 '~Spare WB1[63].6'; 2023 '~Spare WB1[63].7'; 2024 '~Spare WB1[63].8'; 2025 '~Spare WB1[63].9'; 2026 '~Spare WB1[63].10'; 2027 '~Spare WB1[63].11'; 2028 '~Spare WB1[63].12'; 2029 '~Spare WB1[63].13'; 2030 '~Spare WB1[63].14'; 2031 '~Spare WB1[63].15'; 2032 '~Spare WB1[63].16'; 2033 '~Spare WB1[63].17'; 2034 '~Spare WB1[63].18'; 2035 '~Spare WB1[63].19'; 2036 '~Spare WB1[63].20'; 2037 '~Spare WB1[63].21'; 2038 '~Spare WB1[63].22'; 2039 '~Spare WB1[63].23'; 2040 '~Spare WB1[63].24'; 2041 '~Spare WB1[63].25'; 2042 '~Spare WB1[63].26'; 2043 '~Spare WB1[63].27'; 2044 '~Spare WB1[63].28'; 2045 '~Spare WB1[63].29'; 2046 '~Spare WB1[63].30'; 2047 '~Spare WB1[63].31'; 2048 '~Spare WB1[64].0'; 2049 '~Spare WB1[64].1'; 2050 '~Spare WB1[64].2'; 2051 '~Spare WB1[64].3'; 2052 '~Spare WB1[64].4'; 2053 '~Spare WB1[64].5'; 2054 '~Spare WB1[64].6'; 2055 '~Spare WB1[64].7'; 2056 '~Spare WB1[64].8'; 2057 '~Spare WB1[64].9'; 2058 '~Spare WB1[64].10'; 2059 '~Spare WB1[64].11'; 2060 '~Spare WB1[64].12'; 2061 '~Spare WB1[64].13'; 2062 '~Spare WB1[64].14'; 2063 '~Spare WB1[64].15'; 2064 '~Spare WB1[64].16'; 2065 '~Spare WB1[64].17'; 2066 '~Spare WB1[64].18'; 2067 '~Spare WB1[64].19'; 2068 '~Spare WB1[64].20'; 2069 '~Spare WB1[64].21'; 2070 '~Spare WB1[64].22'; 2071 '~Spare WB1[64].23'; 2072 '~Spare WB1[64].24'; 2073 '~Spare WB1[64].25'; 2074 '~Spare WB1[64].26'; 2075 '~Spare WB1[64].27'; 2076 '~Spare WB1[64].28'; 2077 '~Spare WB1[64].29'; 2078 '~Spare WB1[64].30'; 2079 '~Spare WB1[64].31'; 2080 '~Spare WB1[65].0'; 2081 '~Spare WB1[65].1'; 2082 '~Spare WB1[65].2'; 2083 '~Spare WB1[65].3'; 2084 '~Spare WB1[65].4'; 2085 '~Spare WB1[65].5'; 2086 '~Spare WB1[65].6'; 2087 '~Spare WB1[65].7'; 2088 '~Spare WB1[65].8'; 2089 '~Spare WB1[65].9'; 2090 '~Spare WB1[65].10'; 2091 '~Spare WB1[65].11'; 2092 '~Spare WB1[65].12'; 2093 '~Spare WB1[65].13'; 2094 '~Spare WB1[65].14'; 2095 '~Spare WB1[65].15'; 2096 '~Spare WB1[65].16'; 2097 '~Spare WB1[65].17'; 2098 '~Spare WB1[65].18'; 2099 '~Spare WB1[65].19'; 2100 '~Spare WB1[65].20'; 2101 '~Spare WB1[65].21'; 2102 '~Spare WB1[65].22'; 2103 '~Spare WB1[65].23'; 2104 '~Spare WB1[65].24'; 2105 '~Spare WB1[65].25'; 2106 '~Spare WB1[65].26'; 2107 '~Spare WB1[65].27'; 2108 '~Spare WB1[65].28'; 2109 '~Spare WB1[65].29'; 2110 '~Spare WB1[65].30'; 2111 '~Spare WB1[65].31'; 2112 '~S001R08 Waiting Zone #1 Not Clear WB1[66].0'; 2113 '~S001R08 Waiting Zone #2 Not Clear WB1[66].1'; 2114 '~S001R08 Waiting Zone #3 Not Clear WB1[66].2'; 2115 '~S001R08 Waiting Zone #4 Not Clear WB1[66].3'; 2116 '~S001R08 Waiting Zone #5 Not Clear WB1[66].4'; 2117 '~S001R08 Waiting Zone #6 Not Clear WB1[66].5'; 2118 '~S001R08 Waiting Zone #7 Not Clear WB1[66].6'; 2119 '~S001R08 Waiting Zone #8 Not Clear WB1[66].7'; 2120 '~S001R08 Waiting Zone #9 Not Clear WB1[66].8'; 2121 '~S001R08 Waiting Zone #10 Not Clear WB1[66].9'; 2122 '~S001R08 Waiting Zone #11 Not Clear WB1[66].10'; 2123 '~S001R08 Waiting Zone #12 Not Clear WB1[66].11'; 2124 '~S001R08 Waiting Zone #13 Not Clear WB1[66].12'; 2125 '~S001R08 Waiting Zone #14 Not Clear WB1[66].13'; 2126 '~S001R08 Waiting Tip Dress Zone #1 Not Clear WB1[66].14'; 2127 '~S001R08 Waiting Tip Dress Zone #2 Not Clear WB1[66].15'; 2128 '~S001R08 Adjacent Robot xx-xx In Teach WB1[66].16'; 2129 '~S001R08 Adjacent Robot xx-xx In Teach WB1[66].17'; 2130 '~S001R08 Adjacent Robot xx-xx In Teach WB1[66].18'; 2131 '~S001R08 Adjacent Robot xx-xx In Teach WB1[66].19'; 2132 '~S001R08 Adjacent Robot xx-xx In Teach WB1[66].20'; 2133 '~S001R08 Adjacent Robot xx-xx In Teach WB1[66].21'; 2134 '~S001R08 Adjacent Robot xx-xx In Teach WB1[66].22'; 2135 '~S001R08 Adjacent Robot xx-xx In Teach WB1[66].23'; 2136 '~S001R08 Adjacent Robot xx-xx In Teach WB1[66].24'; 2137 '~S001R08 Adjacent Robot xx-xx In Teach WB1[66].25'; 2138 '~Spare WB1[66].26'; 2139 '~Spare WB1[66].27'; 2140 '~Spare WB1[66].28'; 2141 '~S001R08 Robot Not Clear Of Fixture WB1[66].29'; 2142 '~Spare WB1[66].30'; 2143 '~Spare WB1[66].31'; 2144 '~Spare WB1[67].0'; 2145 '~Spare WB1[67].1'; 2146 '~Spare WB1[67].2'; 2147 '~Spare WB1[67].3'; 2148 '~Spare WB1[67].4'; 2149 '~Spare WB1[67].5'; 2150 '~Spare WB1[67].6'; 2151 '~Spare WB1[67].7'; 2152 '~Spare WB1[67].8'; 2153 '~Spare WB1[67].9'; 2154 '~Spare WB1[67].10'; 2155 '~Spare WB1[67].11'; 2156 '~Spare WB1[67].12'; 2157 '~Spare WB1[67].13'; 2158 '~Spare WB1[67].14'; 2159 '~Spare WB1[67].15'; 2160 '~Spare WB1[67].16'; 2161 '~Spare WB1[67].17'; 2162 '~Spare WB1[67].18'; 2163 '~Spare WB1[67].19'; 2164 '~Spare WB1[67].20'; 2165 '~Spare WB1[67].21'; 2166 '~Spare WB1[67].22'; 2167 '~Spare WB1[67].23'; 2168 '~Spare WB1[67].24'; 2169 '~Spare WB1[67].25'; 2170 '~Spare WB1[67].26'; 2171 '~Spare WB1[67].27'; 2172 '~Spare WB1[67].28'; 2173 '~Spare WB1[67].29'; 2174 '~Spare WB1[67].30'; 2175 '~Spare WB1[67].31'; 2176 '~S001R08 Cycle Overtime WB1[68].0'; 2177 '~S001R08 In Bypass WB1[68].1'; 2178 '~S001R08 Battery Low WB1[68].2'; 2179 '~S001R08 Servo Over Torque WB1[68].3'; 2180 '~S001R08 Process Retry In Progress WB1[68].4'; 2181 '~Spare WB1[68].5'; 2182 '~S001R08 Robot Edit Occurred Ext App WB1[68].6'; 2183 '~S001R08 Robot Input Simmed WB1[68].7'; 2184 '~S001R08 Robot Output Simmed WB1[68].8'; 2185 '~Spare WB1[68].9'; 2186 '~Spare WB1[68].10'; 2187 '~Spare WB1[68].11'; 2188 '~Spare WB1[68].12'; 2189 '~Spare WB1[68].13'; 2190 '~Spare WB1[68].14'; 2191 '~Spare WB1[68].15'; 2192 '~S001R08F1B1.M.ModuleFlt - Externa App 1 I/O Module Warning WB1[68].16'; 2193 '~S001R08F2B1.M.ModuleFlt - Externa App 2 I/O Module Warning WB1[68].17'; 2194 '~S001R08F3B1.M.ModuleFlt - Externa App 3 I/O Module Warning WB1[68].18'; 2195 '~Spare WB1[68].19'; 2196 '~Spare WB1[68].20'; 2197 '~Spare WB1[68].21'; 2198 '~Spare WB1[68].22'; 2199 '~Spare WB1[68].23'; 2200 '~S001R08ES1 - S001R08 EtherNet Switch Port At Half Duplex WB1[68].24'; 2201 '~S001R08ES1 - S001R08 EtherNet Switch Config Changes Not Saved WB1[68].25'; 2202 '~S001R08ES1 - S001R08 EtherNet Switch Configuration Changed WB1[68].26'; 2203 '~S001R08ES1 - S001R08 EtherNet Switch Port With Excessive Errors WB1[68].27'; 2204 '~S001R08ES1 - S001R08 EtherNet Switch Port With Utilization Warning WB1[68].28'; 2205 '~S001R08ES1 - S001R08 EtherNet Switch Changes Require Reboot WB1[68].29'; 2206 '~Spare WB1[68].30'; 2207 '~Spare WB1[68].31'; 2208 '~Spare WB1[69].0'; 2209 '~Spare WB1[69].1'; 2210 '~S001R08 Servo Gun Tip Calib Request 1 WB1[69].2'; 2211 '~S001R08 I-Available Warning 1 WB1[69].3'; 2212 '~S001R08 Tip Dress Motor 1 Fault Bypassed WB1[69].4'; 2213 '~S001R08 Tip Change Notice 1 WB1[69].5'; 2214 '~S001R08 Bypass Tip Dresser 1 Selected WB1[69].6'; 2215 '~S001R08 Auto Tip Changer Low 1 WB1[69].7'; 2216 '~S001R08 Auto Tip Changer Empty 1 WB1[69].8'; 2217 '~S001R08 Tip Wear Ratio Warning 1 - Touch Up Tip Dress Program WB1[69].9'; 2218 '~S001R08 Stud Weld 1 Maintenance Reqd WB1[69].10'; 2219 '~S001R08 Stud Weld 1 Low Stud Warning WB1[69].11'; 2220 '~Spare WB1[69].12'; 2221 '~S001R08 Rivet 1 Low Rivet Warning WB1[69].13'; 2222 '~S001R08 Rivet 1 - Skip Once Initiated from Robot TP WB1[69].14'; 2223 '~S001R08 Rivet 1 - Skip Remaining Initiated from Robot TP WB1[69].15'; 2224 '~S001R08 Rivet 1 Preventive Maintenace Required WB1[69].16'; 2225 '~S001R08 Rivet 1 Magazine Low WB1[69].17'; 2226 '~S001R08 Tip Change 1 Bypassed WB1[69].18'; 2227 '~S001R08 Mig Weld Fluid Level Low WB1[69].19'; 2228 '~S001R08 Weld Ctrlr 1 Adaptive Mode Is Disabled WB1[69].20'; 2229 '~S001R08 Tip Cutter 1 Warning WB1[69].21'; 2230 '~S001R08 Rivet 1 Tape-Cut Required WB1[69].22'; 2231 '~S001R08 Wire Feeder Motor Over Current WB1[69].23'; 2232 '~Spare WB1[69].24'; 2233 '~S001R08 Sealer Ctrlr 1 Minor Fault WB1[69].25'; 2234 '~S001R08 Sealer Ctrlr 1 Required Rezeroing WB1[69].26'; 2235 '~S001R08 Loaded To Average WB1[69].27'; 2236 '~S001R08 Vision Process Aborted WB1[69].28'; 2237 '~S001R08 Vision System Trending WB1[69].29'; 2238 '~S001R08 Vision Out Of Tolerance WB1[69].30'; 2239 '~Spare WB1[69].31'; 2240 '~Spare WB1[70].0'; 2241 '~Spare WB1[70].1'; 2242 '~S001R08 Servo Gun Tip Calib Request 2 WB1[70].2'; 2243 '~S001R08 I-Available Warning 2 WB1[70].3'; 2244 '~S001R08 Tip Dress Motor 2 Fault Bypassed WB1[70].4'; 2245 '~S001R08 Tip Change Notice 2 WB1[70].5'; 2246 '~S001R08 Bypass Tip Dresser 2 Selected WB1[70].6'; 2247 '~S001R08 Auto Tip Changer Low 2 WB1[70].7'; 2248 '~S001R08 Auto Tip Changer Empty 2 WB1[70].8'; 2249 '~S001R08 Tip Wear Ratio Warning 2 - Touch Up Tip Dress Program WB1[70].9'; 2250 '~S001R08 Stud Weld 2 Maintenance Reqd WB1[70].10'; 2251 '~S001R08 Stud Weld 2 Low Stud Warning WB1[70].11'; 2252 '~Spare WB1[70].12'; 2253 '~S001R08 Rivet 2 Low Rivet Warning WB1[70].13'; 2254 '~S001R08 Rivet 2 - Skip Once Initiated from Robot TP WB1[70].14'; 2255 '~S001R08 Rivet 2 - Skip Remaining Initiated from Robot TP WB1[70].15'; 2256 '~S001R08 Rivet 2 Preventive Maintenace Required WB1[70].16'; 2257 '~S001R08 Rivet 2 Magazine Low WB1[70].17'; 2258 '~S001R08 Tip Change 2 Bypassed WB1[70].18'; 2259 '~S001R08 Laser Dirty Glass Warning WB1[70].19'; 2260 '~S001R08 Weld Ctrlr 2 Adaptive Mode Is Disabled WB1[70].20'; 2261 '~S001R08 Tip Cutter 2 Warning WB1[70].21'; 2262 '~S001R08 Rivet 2 Tape-Cut Required WB1[70].22'; 2263 '~S001R08 Mig Tip Nozzel Replacement Warning WB1[70].23'; 2264 '~S001R08 Mig Tip Nozzel Replacement Required WB1[70].24'; 2265 '~S001R08 Sealer Ctrlr 2 Minor Fault WB1[70].25'; 2266 '~S001R08 Sealer Ctrlr 2 Required Rezeroing WB1[70].26'; 2267 '~S001R08 Mig Barrel Replacement Warning WB1[70].27'; 2268 '~S001R08 Mig Barrel Replacement Required WB1[70].28'; 2269 '~S001R08 In Touch Up Mode WB1[70].29'; 2270 '~S001R08 Touch Up Mode Not Enabled WB1[70].30'; 2271 '~Spare WB1[70].31'; 2272 '~S001R08 Laser Controller Fault WB1[71].0'; 2273 '~S001R08 Laser Dirty Glass Warning WB1[71].1'; 2274 '~S001R08 Laser Warning WB1[71].2'; 2275 '~Spare WB1[71].3'; 2276 '~Spare WB1[71].4'; 2277 '~Spare WB1[71].5'; 2278 '~Spare WB1[71].6'; 2279 '~Spare WB1[71].7'; 2280 '~Spare WB1[71].8'; 2281 '~Spare WB1[71].9'; 2282 '~Spare WB1[71].10'; 2283 '~Spare WB1[71].11'; 2284 '~Spare WB1[71].12'; 2285 '~Spare WB1[71].13'; 2286 '~Spare WB1[71].14'; 2287 '~Spare WB1[71].15'; 2288 '~Spare WB1[71].16'; 2289 '~Spare WB1[71].17'; 2290 '~Spare WB1[71].18'; 2291 '~Spare WB1[71].19'; 2292 '~Spare WB1[71].20'; 2293 '~Spare WB1[71].21'; 2294 '~Spare WB1[71].22'; 2295 '~Spare WB1[71].23'; 2296 '~Spare WB1[71].24'; 2297 '~Spare WB1[71].25'; 2298 '~Spare WB1[71].26'; 2299 '~Spare WB1[71].27'; 2300 '~Spare WB1[71].28'; 2301 '~Spare WB1[71].29'; 2302 '~Spare WB1[71].30'; 2303 '~Spare WB1[71].31'; 2304 '~Spare WB1[72].0'; 2305 '~Spare WB1[72].1'; 2306 '~Spare WB1[72].2'; 2307 '~Spare WB1[72].3'; 2308 '~Spare WB1[72].4'; 2309 '~Spare WB1[72].5'; 2310 '~Spare WB1[72].6'; 2311 '~Spare WB1[72].7'; 2312 '~Spare WB1[72].8'; 2313 '~Spare WB1[72].9'; 2314 '~Spare WB1[72].10'; 2315 '~Spare WB1[72].11'; 2316 '~Spare WB1[72].12'; 2317 '~Spare WB1[72].13'; 2318 '~Spare WB1[72].14'; 2319 '~Spare WB1[72].15'; 2320 '~Spare WB1[72].16'; 2321 '~Spare WB1[72].17'; 2322 '~Spare WB1[72].18'; 2323 '~Spare WB1[72].19'; 2324 '~Spare WB1[72].20'; 2325 '~Spare WB1[72].21'; 2326 '~Spare WB1[72].22'; 2327 '~Spare WB1[72].23'; 2328 '~Spare WB1[72].24'; 2329 '~Spare WB1[72].25'; 2330 '~Spare WB1[72].26'; 2331 '~Spare WB1[72].27'; 2332 '~Spare WB1[72].28'; 2333 '~Spare WB1[72].29'; 2334 '~Spare WB1[72].30'; 2335 '~Spare WB1[72].31'; 2336 '~Spare WB1[73].0'; 2337 '~Spare WB1[73].1'; 2338 '~Spare WB1[73].2'; 2339 '~Spare WB1[73].3'; 2340 '~Spare WB1[73].4'; 2341 '~Spare WB1[73].5'; 2342 '~Spare WB1[73].6'; 2343 '~Spare WB1[73].7'; 2344 '~Spare WB1[73].8'; 2345 '~Spare WB1[73].9'; 2346 '~Spare WB1[73].10'; 2347 '~Spare WB1[73].11'; 2348 '~Spare WB1[73].12'; 2349 '~Spare WB1[73].13'; 2350 '~Spare WB1[73].14'; 2351 '~Spare WB1[73].15'; 2352 '~Spare WB1[73].16'; 2353 '~Spare WB1[73].17'; 2354 '~Spare WB1[73].18'; 2355 '~Spare WB1[73].19'; 2356 '~Spare WB1[73].20'; 2357 '~Spare WB1[73].21'; 2358 '~Spare WB1[73].22'; 2359 '~Spare WB1[73].23'; 2360 '~Spare WB1[73].24'; 2361 '~Spare WB1[73].25'; 2362 '~Spare WB1[73].26'; 2363 '~Spare WB1[73].27'; 2364 '~Spare WB1[73].28'; 2365 '~Spare WB1[73].29'; 2366 '~Spare WB1[73].30'; 2367 '~Spare WB1[73].31'; 2368 '~Spare WB1[74].0'; 2369 '~Spare WB1[74].1'; 2370 '~Spare WB1[74].2'; 2371 '~Spare WB1[74].3'; 2372 '~Spare WB1[74].4'; 2373 '~Spare WB1[74].5'; 2374 '~Spare WB1[74].6'; 2375 '~Spare WB1[74].7'; 2376 '~Spare WB1[74].8'; 2377 '~Spare WB1[74].9'; 2378 '~Spare WB1[74].10'; 2379 '~Spare WB1[74].11'; 2380 '~Spare WB1[74].12'; 2381 '~Spare WB1[74].13'; 2382 '~Spare WB1[74].14'; 2383 '~Spare WB1[74].15'; 2384 '~Spare WB1[74].16'; 2385 '~Spare WB1[74].17'; 2386 '~Spare WB1[74].18'; 2387 '~Spare WB1[74].19'; 2388 '~Spare WB1[74].20'; 2389 '~Spare WB1[74].21'; 2390 '~Spare WB1[74].22'; 2391 '~Spare WB1[74].23'; 2392 '~Spare WB1[74].24'; 2393 '~Spare WB1[74].25'; 2394 '~Spare WB1[74].26'; 2395 '~Spare WB1[74].27'; 2396 '~Spare WB1[74].28'; 2397 '~Spare WB1[74].29'; 2398 '~Spare WB1[74].30'; 2399 '~Spare WB1[74].31'; 2400 '~S001 Fixture Cycle Over Time WB1[75].0'; 2401 '~Spare WB1[75].1'; 2402 '~Spare WB1[75].2'; 2403 '~Spare WB1[75].3'; 2404 '~Spare WB1[75].4'; 2405 '~Spare WB1[75].5'; 2406 '~Spare WB1[75].6'; 2407 '~Spare WB1[75].7'; 2408 '~Spare WB1[75].8'; 2409 '~Spare WB1[75].9'; 2410 '~Spare WB1[75].10'; 2411 '~Spare WB1[75].11'; 2412 '~Spare WB1[75].12'; 2413 '~Spare WB1[75].13'; 2414 '~Spare WB1[75].14'; 2415 '~Spare WB1[75].15'; 2416 '~Spare WB1[75].16'; 2417 '~Spare WB1[75].17'; 2418 '~Spare WB1[75].18'; 2419 '~Spare WB1[75].19'; 2420 '~Spare WB1[75].20'; 2421 '~Spare WB1[75].21'; 2422 '~Spare WB1[75].22'; 2423 '~Spare WB1[75].23'; 2424 '~Spare WB1[75].24'; 2425 '~Spare WB1[75].25'; 2426 '~Spare WB1[75].26'; 2427 '~Spare WB1[75].27'; 2428 '~Spare WB1[75].28'; 2429 '~Spare WB1[75].29'; 2430 '~Spare WB1[75].30'; 2431 '~Spare WB1[75].31'; 2432 '~Spare WB1[76].0'; 2433 '~Spare WB1[76].1'; 2434 '~Spare WB1[76].2'; 2435 '~Spare WB1[76].3'; 2436 '~Spare WB1[76].4'; 2437 '~Spare WB1[76].5'; 2438 '~Spare WB1[76].6'; 2439 '~Spare WB1[76].7'; 2440 '~Spare WB1[76].8'; 2441 '~Spare WB1[76].9'; 2442 '~Spare WB1[76].10'; 2443 '~Spare WB1[76].11'; 2444 '~Spare WB1[76].12'; 2445 '~Spare WB1[76].13'; 2446 '~Spare WB1[76].14'; 2447 '~Spare WB1[76].15'; 2448 '~Spare WB1[76].16'; 2449 '~Spare WB1[76].17'; 2450 '~Spare WB1[76].18'; 2451 '~Spare WB1[76].19'; 2452 '~Spare WB1[76].20'; 2453 '~Spare WB1[76].21'; 2454 '~Spare WB1[76].22'; 2455 '~Spare WB1[76].23'; 2456 '~Spare WB1[76].24'; 2457 '~Spare WB1[76].25'; 2458 '~Spare WB1[76].26'; 2459 '~Spare WB1[76].27'; 2460 '~Spare WB1[76].28'; 2461 '~Spare WB1[76].29'; 2462 '~Spare WB1[76].30'; 2463 '~Spare WB1[76].31'; 2464 '~Spare WB1[77].0'; 2465 '~Spare WB1[77].1'; 2466 '~Spare WB1[77].2'; 2467 '~Spare WB1[77].3'; 2468 '~Spare WB1[77].4'; 2469 '~Spare WB1[77].5'; 2470 '~Spare WB1[77].6'; 2471 '~Spare WB1[77].7'; 2472 '~Spare WB1[77].8'; 2473 '~Spare WB1[77].9'; 2474 '~Spare WB1[77].10'; 2475 '~Spare WB1[77].11'; 2476 '~Spare WB1[77].12'; 2477 '~Spare WB1[77].13'; 2478 '~Spare WB1[77].14'; 2479 '~Spare WB1[77].15'; 2480 '~Spare WB1[77].16'; 2481 '~Spare WB1[77].17'; 2482 '~Spare WB1[77].18'; 2483 '~Spare WB1[77].19'; 2484 '~Spare WB1[77].20'; 2485 '~Spare WB1[77].21'; 2486 '~Spare WB1[77].22'; 2487 '~Spare WB1[77].23'; 2488 '~Spare WB1[77].24'; 2489 '~Spare WB1[77].25'; 2490 '~Spare WB1[77].26'; 2491 '~Spare WB1[77].27'; 2492 '~Spare WB1[77].28'; 2493 '~Spare WB1[77].29'; 2494 '~Spare WB1[77].30'; 2495 '~Spare WB1[77].31'; 2496 '~Spare WB1[78].0'; 2497 '~Spare WB1[78].1'; 2498 '~Spare WB1[78].2'; 2499 '~Spare WB1[78].3'; 2500 '~Spare WB1[78].4'; 2501 '~Spare WB1[78].5'; 2502 '~Spare WB1[78].6'; 2503 '~Spare WB1[78].7'; 2504 '~Spare WB1[78].8'; 2505 '~Spare WB1[78].9'; 2506 '~Spare WB1[78].10'; 2507 '~Spare WB1[78].11'; 2508 '~Spare WB1[78].12'; 2509 '~Spare WB1[78].13'; 2510 '~Spare WB1[78].14'; 2511 '~Spare WB1[78].15'; 2512 '~Spare WB1[78].16'; 2513 '~Spare WB1[78].17'; 2514 '~Spare WB1[78].18'; 2515 '~Spare WB1[78].19'; 2516 '~Spare WB1[78].20'; 2517 '~Spare WB1[78].21'; 2518 '~Spare WB1[78].22'; 2519 '~Spare WB1[78].23'; 2520 '~Spare WB1[78].24'; 2521 '~Spare WB1[78].25'; 2522 '~Spare WB1[78].26'; 2523 '~Spare WB1[78].27'; 2524 '~Spare WB1[78].28'; 2525 '~Spare WB1[78].29'; 2526 '~Spare WB1[78].30'; 2527 '~Spare WB1[78].31'; 2528 '~Spare WB1[79].0'; 2529 '~Spare WB1[79].1'; 2530 '~Spare WB1[79].2'; 2531 '~Spare WB1[79].3'; 2532 '~Spare WB1[79].4'; 2533 '~Spare WB1[79].5'; 2534 '~Spare WB1[79].6'; 2535 '~Spare WB1[79].7'; 2536 '~Spare WB1[79].8'; 2537 '~Spare WB1[79].9'; 2538 '~Spare WB1[79].10'; 2539 '~Spare WB1[79].11'; 2540 '~Spare WB1[79].12'; 2541 '~Spare WB1[79].13'; 2542 '~Spare WB1[79].14'; 2543 '~Spare WB1[79].15'; 2544 '~Spare WB1[79].16'; 2545 '~Spare WB1[79].17'; 2546 '~Spare WB1[79].18'; 2547 '~Spare WB1[79].19'; 2548 '~Spare WB1[79].20'; 2549 '~Spare WB1[79].21'; 2550 '~Spare WB1[79].22'; 2551 '~Spare WB1[79].23'; 2552 '~Spare WB1[79].24'; 2553 '~Spare WB1[79].25'; 2554 '~Spare WB1[79].26'; 2555 '~Spare WB1[79].27'; 2556 '~Spare WB1[79].28'; 2557 '~Spare WB1[79].29'; 2558 '~Spare WB1[79].30'; 2559 '~Spare WB1[79].31'; 2560 '~Spare WB1[80].0'; 2561 '~Spare WB1[80].1'; 2562 '~Spare WB1[80].2'; 2563 '~Spare WB1[80].3'; 2564 '~Spare WB1[80].4'; 2565 '~Spare WB1[80].5'; 2566 '~Spare WB1[80].6'; 2567 '~Spare WB1[80].7'; 2568 '~Spare WB1[80].8'; 2569 '~Spare WB1[80].9'; 2570 '~Spare WB1[80].10'; 2571 '~Spare WB1[80].11'; 2572 '~Spare WB1[80].12'; 2573 '~Spare WB1[80].13'; 2574 '~Spare WB1[80].14'; 2575 '~Spare WB1[80].15'; 2576 '~Spare WB1[80].16'; 2577 '~Spare WB1[80].17'; 2578 '~Spare WB1[80].18'; 2579 '~Spare WB1[80].19'; 2580 '~Spare WB1[80].20'; 2581 '~Spare WB1[80].21'; 2582 '~Spare WB1[80].22'; 2583 '~Spare WB1[80].23'; 2584 '~Spare WB1[80].24'; 2585 '~Spare WB1[80].25'; 2586 '~Spare WB1[80].26'; 2587 '~Spare WB1[80].27'; 2588 '~Spare WB1[80].28'; 2589 '~Spare WB1[80].29'; 2590 '~Spare WB1[80].30'; 2591 '~Spare WB1[80].31'; 2592 '~Spare WB1[81].0'; 2593 '~Spare WB1[81].1'; 2594 '~Spare WB1[81].2'; 2595 '~Spare WB1[81].3'; 2596 '~Spare WB1[81].4'; 2597 '~Spare WB1[81].5'; 2598 '~Spare WB1[81].6'; 2599 '~Spare WB1[81].7'; 2600 '~Spare WB1[81].8'; 2601 '~Spare WB1[81].9'; 2602 '~Spare WB1[81].10'; 2603 '~Spare WB1[81].11'; 2604 '~Spare WB1[81].12'; 2605 '~Spare WB1[81].13'; 2606 '~Spare WB1[81].14'; 2607 '~Spare WB1[81].15'; 2608 '~Spare WB1[81].16'; 2609 '~Spare WB1[81].17'; 2610 '~Spare WB1[81].18'; 2611 '~Spare WB1[81].19'; 2612 '~Spare WB1[81].20'; 2613 '~Spare WB1[81].21'; 2614 '~Spare WB1[81].22'; 2615 '~Spare WB1[81].23'; 2616 '~Spare WB1[81].24'; 2617 '~Spare WB1[81].25'; 2618 '~Spare WB1[81].26'; 2619 '~Spare WB1[81].27'; 2620 '~Spare WB1[81].28'; 2621 '~Spare WB1[81].29'; 2622 '~Spare WB1[81].30'; 2623 '~Spare WB1[81].31'; 2624 '~Spare WB1[82].0'; 2625 '~Spare WB1[82].1'; 2626 '~Spare WB1[82].2'; 2627 '~Spare WB1[82].3'; 2628 '~Spare WB1[82].4'; 2629 '~Spare WB1[82].5'; 2630 '~Spare WB1[82].6'; 2631 '~Spare WB1[82].7'; 2632 '~Spare WB1[82].8'; 2633 '~Spare WB1[82].9'; 2634 '~Spare WB1[82].10'; 2635 '~Spare WB1[82].11'; 2636 '~Spare WB1[82].12'; 2637 '~Spare WB1[82].13'; 2638 '~Spare WB1[82].14'; 2639 '~Spare WB1[82].15'; 2640 '~Spare WB1[82].16'; 2641 '~Spare WB1[82].17'; 2642 '~Spare WB1[82].18'; 2643 '~Spare WB1[82].19'; 2644 '~Spare WB1[82].20'; 2645 '~Spare WB1[82].21'; 2646 '~Spare WB1[82].22'; 2647 '~Spare WB1[82].23'; 2648 '~Spare WB1[82].24'; 2649 '~Spare WB1[82].25'; 2650 '~Spare WB1[82].26'; 2651 '~Spare WB1[82].27'; 2652 '~Spare WB1[82].28'; 2653 '~Spare WB1[82].29'; 2654 '~Spare WB1[82].30'; 2655 '~Spare WB1[82].31'; 2656 '~Spare WB1[83].0'; 2657 '~Spare WB1[83].1'; 2658 '~Spare WB1[83].2'; 2659 '~Spare WB1[83].3'; 2660 '~Spare WB1[83].4'; 2661 '~Spare WB1[83].5'; 2662 '~Spare WB1[83].6'; 2663 '~Spare WB1[83].7'; 2664 '~Spare WB1[83].8'; 2665 '~Spare WB1[83].9'; 2666 '~Spare WB1[83].10'; 2667 '~Spare WB1[83].11'; 2668 '~Spare WB1[83].12'; 2669 '~Spare WB1[83].13'; 2670 '~Spare WB1[83].14'; 2671 '~Spare WB1[83].15'; 